// TIA Portal project "Urban Intersection Control System" (V17)

(* hardware
DEVICE "S7-1500/ET200MP station_1"  S7-1500 station
   slot 0: "Rail_0"  Rack  6ES7 590-1***0-0AA0
   slot 1: "PLC_UICS_01"  CPU 1512C-1 PN  6ES7 512-1CK00-0AB0  V2.9
      slot 3: "CPU display_1"  6ES7591-1AA00-0AA0
      slot 32768: "PROFINET interface_1"  X1
         slot 32769: "Port_1"  X1 P1
         slot 32770: "Port_2"  X1 P2
      slot 34817: "Virtual CP interface port_1"  Virtual CP interface port  Virtual CP interface port
DEVICE "HMI_1"  KTP1200 Basic PN
   slot 0: "HMI_1"  KTP1200 Basic PN  6AV2 123-2MB03-0AX0  17.0.0.0
   slot 1: "HMI_RT_1"  KTP1200 Basic PN  6AV2 123-2MB03-0AX0  17.0.0.0
   slot 5: "HMI_1.IE_CP_1"  PROFINET Interface  17.0.0.0
      slot 1: "PROFINET Interface_1"  PROFINET Interface
         slot 1: "Port_1"  Port
*)

// ===== PLC "PLC_UICS_01"  CPU 1512C-1 PN =====

VAR_GLOBAL   // PLC tag table "UICS_Table"
   "PB_Ped_Main_East" AT %I10.2 : Bool;   // Push button for pedestrian crossing on eastern Main Street
   "PB_Ped_Main_West" AT %I10.3 : Bool;   // Push button for pedestrian crossing on western Main Street
   "EM_Main_Override" AT %I10.6 : Bool;   // Emergency override signal (e.g. ambulances) on Main Street
   "EM_Cross_Override" AT %I10.7 : Bool;   // Emergency override signal on Cross Street
   "SENSOR_Main_Vehicle" AT %I11.0 : Bool;   // Vehicle detection sensor on Main Street
   "SENSOR_Cross_Vehicle" AT %I11.1 : Bool;   // Vehicle detection sensor on Cross Street
   "TL_Main_Red_West" AT %Q4.0 : Bool;   // Red traffic light signal for western Main Street
   "TL_Main_Yellow_West" AT %Q4.2 : Bool;   // Yellow traffic light signal for western Main Street
   "TL_Main_Green_West" AT %Q4.4 : Bool;   // Green traffic light signal for western Main Street
   "TL_Cross_Red_North" AT %Q4.6 : Bool;   // Red traffic light signal for northern Cross Street
   "TL_Cross_Yellow_North" AT %Q5.0 : Bool;   // Yellow traffic light signal for northern Cross Street
   "TL_Cross_Green_North" AT %Q5.2 : Bool;   // Green traffic light signal for northern Cross Street
   "PED_Main_Walk_West" AT %Q5.4 : Bool;   // Pedestrian walk signal for western Main Street
   "PED_Main_DontWalk_West" AT %Q5.6 : Bool;   // Pedestrian don’t-walk signal for western Main Street
   "PED_Cross_Walk_North" AT %Q6.0 : Bool;   // Pedestrian walk signal for northern Cross Street
   "PED_Cross_DontWalk_North" AT %Q6.2 : Bool;   // Pedestrian don’t-walk signal for northern Cross Street
   "PED_Warning_Buzzer" AT %Q6.4 : Bool;   // Audible alert for pedestrian crossing
   "SYS_Stop" AT %I10.1 : Bool;   // Emergency stop function
   "SYS_Start" AT %I10.0 : Bool;   // Begins the system
   "TL_Main_Red_East" AT %Q4.1 : Bool;   // Red traffic light signal for eastern Main Street
   "TL_Main_Yellow_East" AT %Q4.3 : Bool;   // Yellow traffic light signal for eastern Main Street
   "TL_Main_Green_East" AT %Q4.5 : Bool;   // Green traffic light signal for eastern Main Street
   "TL_Cross_Red_South" AT %Q4.7 : Bool;   // Red traffic light signal for southern Cross Street
   "TL_Cross_Yellow_South" AT %Q5.1 : Bool;   // Yellow traffic light signal for southern Cross Street
   "TL_Cross_Green_South" AT %Q5.3 : Bool;   // Green traffic light signal for southern Cross Street
   "PED_Main_Walk_East" AT %Q5.5 : Bool;   // Pedestrian walk signal for eastern Main Street
   "PED_Main_DontWalk_East" AT %Q5.7 : Bool;   // Pedestrian don’t-walk signal for eastern Main Street
   "PED_Cross_Walk_South" AT %Q6.1 : Bool;   // Pedestrian walk signal for southern Cross Street
   "PED_Cross_DontWalk_South" AT %Q6.3 : Bool;   // Pedestrian don’t-walk signal for southern Cross Street
   "PB_Ped_Cross_South" AT %I10.4 : Bool;   // Push button for pedestrian crossing on southern Cross Street
   "PB_Ped_Cross_North" AT %I10.5 : Bool;   // Push button for pedestrian crossing on northern Cross Street
   "PED_Main_Queue_East" AT %Q6.5 : Bool;   // Pedestrian queue signal for eastern Main Street
   "PED_Main_Queue_West" AT %Q6.6 : Bool;   // Pedestrian queue signal for western Main Street
   "PED_Cross_Queue_North" AT %Q6.7 : Bool;   // Pedestrian queue signal for southern Cross Street
   "PED_Cross_Queue_South" AT %Q7.0 : Bool;   // Pedestrian queue signal for northern Cross Street
END_VAR

DATA_BLOCK "Main_Control_System_DB"   // DB1
{ S7_Optimized_Access := 'TRUE' }
VERSION : 0.1
// stored: InstanceOfName Main_Control_System
"Main_Control_System"
BEGIN
END_DATA_BLOCK

DATA_BLOCK "Traffic_Light_Operations_DB"   // DB3
{ S7_Optimized_Access := 'TRUE' }
VERSION : 0.1
// stored: InstanceOfName Traffic_Light_Operations
"Traffic_Light_Operations"
BEGIN
END_DATA_BLOCK

DATA_BLOCK "Status_Reset_DB"   // DB7
{ S7_Optimized_Access := 'TRUE' }
VERSION : 0.1
// stored: InstanceOfName Status_Reset
"Status_Reset"
BEGIN
END_DATA_BLOCK

DATA_BLOCK "Pedestrian_Operations_DB"   // DB8
{ S7_Optimized_Access := 'TRUE' }
VERSION : 0.1
// stored: InstanceOfName Pedestrian_Operations
"Pedestrian_Operations"
BEGIN
END_DATA_BLOCK

DATA_BLOCK "Pedestrian_Crossing_DB"   // DB13
{ S7_Optimized_Access := 'TRUE' }
VERSION : 0.1
// stored: InstanceOfName Pedestrian_Crossing
"Pedestrian_Crossing"
BEGIN
END_DATA_BLOCK

// folder: System blocks/Program resources

DATA_BLOCK "MainStEast_Timer_DB"   // DB2
{ S7_Optimized_Access := 'TRUE' }
AUTHOR : Simatic
FAMILY : IEC
NAME : IEC_TMR
VERSION : 1.0
// stored: InstanceOfName IEC_TIMER
"IEC_TIMER"
BEGIN
END_DATA_BLOCK

DATA_BLOCK "CrossStNorth_Timer_DB"   // DB4
{ S7_Optimized_Access := 'TRUE' }
AUTHOR : Simatic
FAMILY : IEC
NAME : IEC_TMR
VERSION : 1.0
// stored: InstanceOfName IEC_TIMER
"IEC_TIMER"
BEGIN
END_DATA_BLOCK

DATA_BLOCK "CrossStSouth_Timer_DB"   // DB5
{ S7_Optimized_Access := 'TRUE' }
AUTHOR : Simatic
FAMILY : IEC
NAME : IEC_TMR
VERSION : 1.0
// stored: InstanceOfName IEC_TIMER
"IEC_TIMER"
BEGIN
END_DATA_BLOCK

DATA_BLOCK "MainStWest_Timer_DB"   // DB6
{ S7_Optimized_Access := 'TRUE' }
AUTHOR : Simatic
FAMILY : IEC
NAME : IEC_TMR
VERSION : 1.0
// stored: InstanceOfName IEC_TIMER
"IEC_TIMER"
BEGIN
END_DATA_BLOCK

DATA_BLOCK "Ped_MainStEast_Timer_DB"   // DB9
{ S7_Optimized_Access := 'TRUE' }
AUTHOR : Simatic
FAMILY : IEC
NAME : IEC_TMR
VERSION : 1.0
// stored: InstanceOfName IEC_TIMER
"IEC_TIMER"
BEGIN
END_DATA_BLOCK

DATA_BLOCK "Ped_MainStWest_Timer_DB"   // DB10
{ S7_Optimized_Access := 'TRUE' }
AUTHOR : Simatic
FAMILY : IEC
NAME : IEC_TMR
VERSION : 1.0
// stored: InstanceOfName IEC_TIMER
"IEC_TIMER"
BEGIN
END_DATA_BLOCK

DATA_BLOCK "Ped_CrossStSouth_Timer_DB"   // DB11
{ S7_Optimized_Access := 'TRUE' }
AUTHOR : Simatic
FAMILY : IEC
NAME : IEC_TMR
VERSION : 1.0
// stored: InstanceOfName IEC_TIMER
"IEC_TIMER"
BEGIN
END_DATA_BLOCK

DATA_BLOCK "Ped_CrossStNorth_Timer_DB"   // DB12
{ S7_Optimized_Access := 'TRUE' }
AUTHOR : Simatic
FAMILY : IEC
NAME : IEC_TMR
VERSION : 1.0
// stored: InstanceOfName IEC_TIMER
"IEC_TIMER"
BEGIN
END_DATA_BLOCK

// folder: (top level)

FUNCTION_BLOCK "Main_Control_System"   // FB1, LAD
{ S7_Optimized_Access := 'TRUE' }
VERSION : 0.1
   VAR_INPUT
      System_Start : Bool;   // Activates the system
      System_Stop : Bool;   // Emergency stop function
   END_VAR
   VAR
      System_Latch : Bool;   // Allows the system to remain active after initially starting up
      System_Running : Bool;   // System is actively running
      Emergency_Stop : Bool;   // Emergency stop activated flag
      HMI_Start_Command : Bool;   // Allows HMI to start the system
      HMI_Stop_Command : Bool;   // Allows HMI to stop the system
      HMI_Latch_Command : Bool;   // Allows HMI visualization to remain active after initially starting up
      HMI_Run_Command : Bool;   // Allows HMI to run the system
   END_VAR
BEGIN

REGION Network 1: System Start
   // Starts the system if all conditions are met
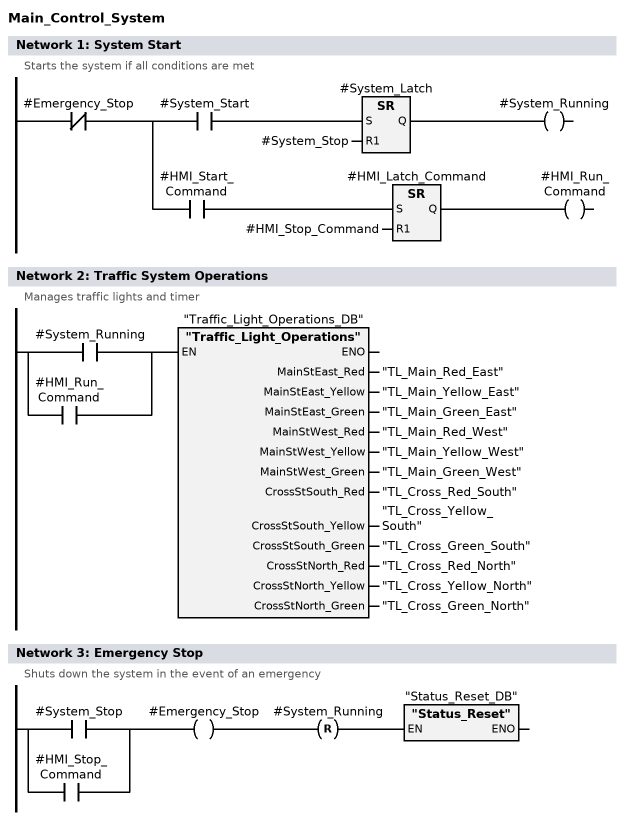
   RUNG wire#powerrail
      I_Contact( #Emergency_Stop )
      wire#w1
      Contact( #System_Start )
      S_SR(operand := #System_Latch, r1 := #System_Stop)
      Coil( #System_Running )
   END_RUNG
   RUNG wire#w1
      Contact( #HMI_Start_Command )
      S_SR(operand := #HMI_Latch_Command, r1 := #HMI_Stop_Command)
      Coil( #HMI_Run_Command )
   END_RUNG
   // the same network as SCL:
   IF NOT #Emergency_Stop AND #System_Start THEN
       #System_Latch := TRUE;   // SR flip-flop
   END_IF;
   IF #System_Stop THEN #System_Latch := FALSE; END_IF;
   #System_Running := #System_Latch;
   IF NOT #Emergency_Stop AND #HMI_Start_Command THEN
       #HMI_Latch_Command := TRUE;   // SR flip-flop
   END_IF;
   IF #HMI_Stop_Command THEN #HMI_Latch_Command := FALSE; END_IF;
   #HMI_Run_Command := #HMI_Latch_Command;
END_REGION

REGION Network 2: Traffic System Operations
   // Manages traffic lights and timer
   RUNG wire#powerrail
      Contact( #System_Running )
      wire#w1
      "Traffic_Light_Operations_DB"(MainStEast_Red => "TL_Main_Red_East", MainStEast_Yellow => "TL_Main_Yellow_East", MainStEast_Green => "TL_Main_Green_East", MainStWest_Red => "TL_Main_Red_West", MainStWest_Yellow => "TL_Main_Yellow_West", MainStWest_Green => "TL_Main_Green_West", CrossStSouth_Red => "TL_Cross_Red_South", CrossStSouth_Yellow => "TL_Cross_Yellow_South", CrossStSouth_Green => "TL_Cross_Green_South", CrossStNorth_Red => "TL_Cross_Red_North", CrossStNorth_Yellow => "TL_Cross_Yellow_North", CrossStNorth_Green => "TL_Cross_Green_North")
   END_RUNG
   RUNG wire#powerrail
      Contact( #HMI_Run_Command )
   END_RUNG wire#w1
   // the same network as SCL:
   IF #System_Running OR #HMI_Run_Command THEN
       "Traffic_Light_Operations_DB"(MainStEast_Red => "TL_Main_Red_East",   // "Traffic_Light_Operations"
                               MainStEast_Yellow => "TL_Main_Yellow_East",
                               MainStEast_Green => "TL_Main_Green_East",
                               MainStWest_Red => "TL_Main_Red_West",
                               MainStWest_Yellow => "TL_Main_Yellow_West",
                               MainStWest_Green => "TL_Main_Green_West",
                               CrossStSouth_Red => "TL_Cross_Red_South",
                               CrossStSouth_Yellow => "TL_Cross_Yellow_South",
                               CrossStSouth_Green => "TL_Cross_Green_South",
                               CrossStNorth_Red => "TL_Cross_Red_North",
                               CrossStNorth_Yellow => "TL_Cross_Yellow_North",
                               CrossStNorth_Green => "TL_Cross_Green_North");
   END_IF;
END_REGION

REGION Network 3: Emergency Stop
   // Shuts down the system in the event of an emergency
   RUNG wire#powerrail
      Contact( #System_Stop )
      wire#w1
      Coil( #Emergency_Stop )
      R_Coil( #System_Running )
      "Status_Reset_DB"()
   END_RUNG
   RUNG wire#powerrail
      Contact( #HMI_Stop_Command )
   END_RUNG wire#w1
   // the same network as SCL:
   #Emergency_Stop := #System_Stop OR #HMI_Stop_Command;
   IF #Emergency_Stop THEN
       #System_Running := FALSE;
       "Status_Reset_DB"();   // "Status_Reset"
   END_IF;
END_REGION
END_FUNCTION_BLOCK

FUNCTION_BLOCK "Traffic_Light_Operations"   // FB2, LAD
{ S7_Optimized_Access := 'TRUE' }
VERSION : 0.1
   VAR_OUTPUT
      MainStEast_Red : Bool;   // Red traffic light signal for eastern Main Street
      MainStEast_Yellow : Bool;   // Yellow traffic light signal for eastern Main Street
      MainStEast_Green : Bool;   // Green traffic light signal for eastern Main Street
      MainStWest_Red : Bool;   // Red traffic light signal for western Main Street
      MainStWest_Yellow : Bool;   // Yellow traffic light signal for western Main Street
      MainStWest_Green : Bool;   // Green traffic light signal for western Main Street
      CrossStSouth_Red : Bool;   // Red traffic light signal for southern Cross Street
      CrossStSouth_Yellow : Bool;   // Yellow traffic light signal for southern Cross Street
      CrossStSouth_Green : Bool;   // Green traffic light signal for southern Cross Street
      CrossStNorth_Red : Bool;   // Red traffic light signal for northern Cross Street
      CrossStNorth_Yellow : Bool;   // Yellow traffic light signal for northern Cross Street
      CrossStNorth_Green : Bool;   // Green traffic light signal for northern Cross Street
   END_VAR
   VAR
      Traffic_Operations_Step : Int;   // Controls the state of traffic operations
      MainStEast_Seconds : Int;   // Allows HMI to read eastern Main Street traffic time
      MainStWest_Seconds : Int;   // Allows HMI to read western Main Street traffic time
      CrossStNorth_Seconds : Int;   // Allows HMI to read northern Cross Street traffic time
      CrossStSouth_Seconds : Int;   // Allows HMI to read southern Cross Street traffic time
      Initialize_Operation : Bool;   // Initiates traffic operations
   END_VAR
   VAR_TEMP
      MainStEast_ET_DInt : DInt;
      MainStEast_ET_Div : DInt;
      CrossStSouth_ET_DInt : DInt;
      CrossStSouth_ET_Div : DInt;
      MainStWest_ET_DInt : DInt;
      MainStWest_ET_Div : DInt;
      CrossStNorth_ET_DInt : DInt;
      CrossStNorth_ET_Div : DInt;
   END_VAR
   VAR_TEMP   // added for the SCL form of the ladder/FBD networks
      _w1 : Bool;
   END_VAR
BEGIN

REGION Network 1: Red Light Control
   // Organization of red traffic lights for Main Street and Cross Street
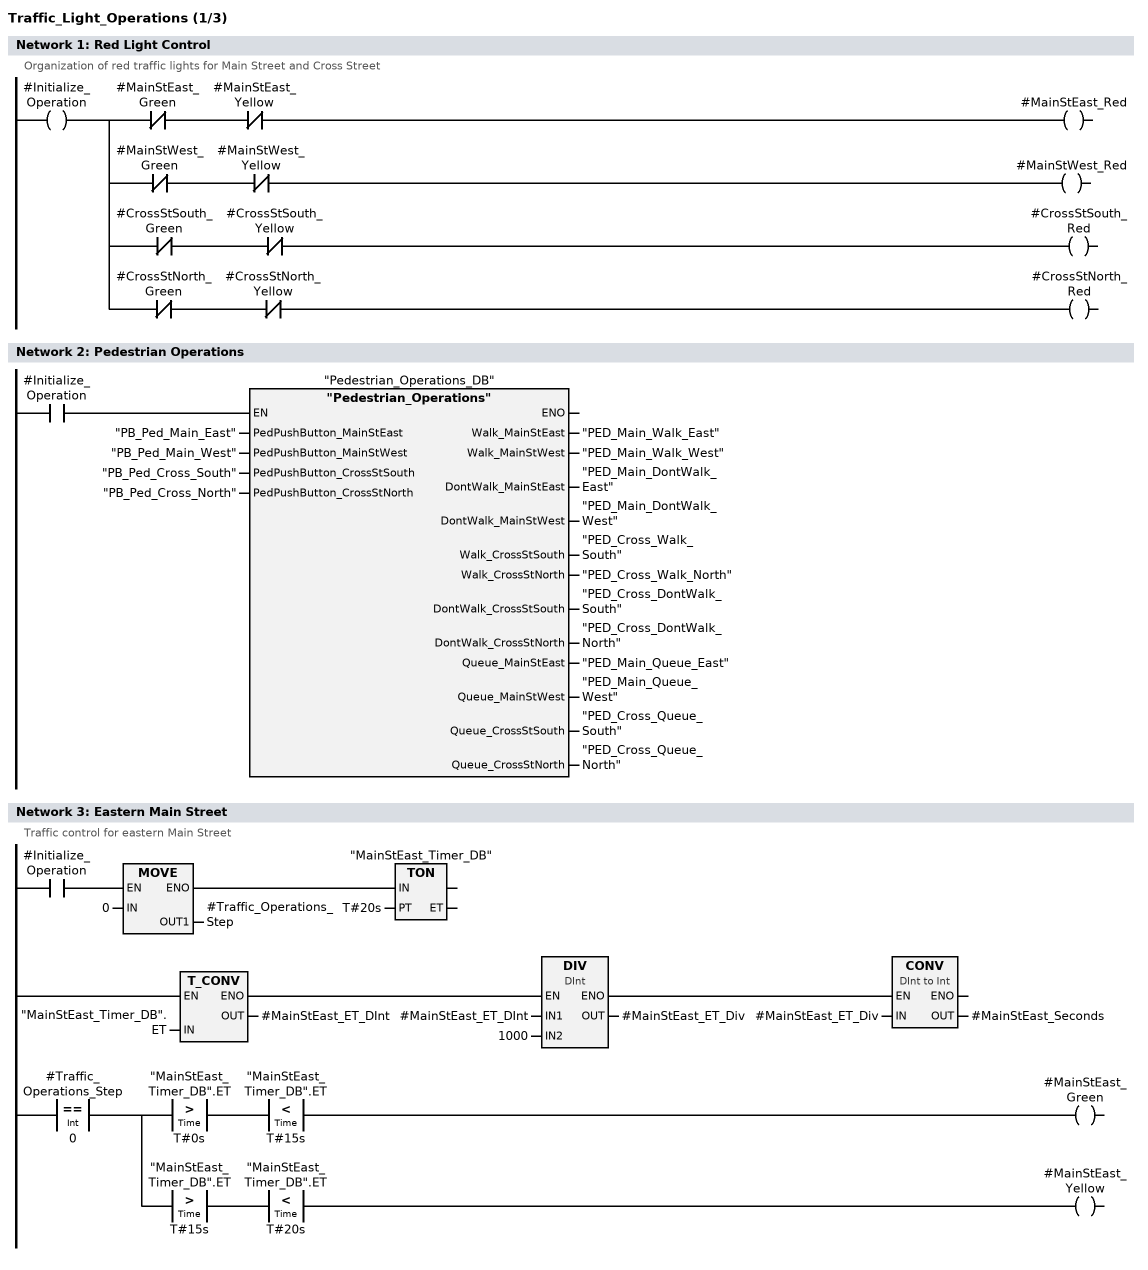
   RUNG wire#powerrail
      Coil( #Initialize_Operation )
      wire#w1
      I_Contact( #MainStEast_Green )
      I_Contact( #MainStEast_Yellow )
      Coil( #MainStEast_Red )
   END_RUNG
   RUNG wire#w1
      I_Contact( #MainStWest_Green )
      I_Contact( #MainStWest_Yellow )
      Coil( #MainStWest_Red )
   END_RUNG
   RUNG wire#w1
      I_Contact( #CrossStSouth_Green )
      I_Contact( #CrossStSouth_Yellow )
      Coil( #CrossStSouth_Red )
   END_RUNG
   RUNG wire#w1
      I_Contact( #CrossStNorth_Green )
      I_Contact( #CrossStNorth_Yellow )
      Coil( #CrossStNorth_Red )
   END_RUNG
   // the same network as SCL:
   #Initialize_Operation := TRUE;
   #MainStEast_Red := NOT #MainStEast_Green AND NOT #MainStEast_Yellow;
   #MainStWest_Red := NOT #MainStWest_Green AND NOT #MainStWest_Yellow;
   #CrossStSouth_Red := NOT #CrossStSouth_Green AND NOT #CrossStSouth_Yellow;
   #CrossStNorth_Red := NOT #CrossStNorth_Green AND NOT #CrossStNorth_Yellow;
END_REGION

REGION Network 2: Pedestrian Operations
   RUNG wire#powerrail
      Contact( #Initialize_Operation )
      "Pedestrian_Operations_DB"(PedPushButton_MainStEast := "PB_Ped_Main_East", PedPushButton_MainStWest := "PB_Ped_Main_West", PedPushButton_CrossStSouth := "PB_Ped_Cross_South", PedPushButton_CrossStNorth := "PB_Ped_Cross_North", Walk_MainStEast => "PED_Main_Walk_East", Walk_MainStWest => "PED_Main_Walk_West", DontWalk_MainStEast => "PED_Main_DontWalk_East", DontWalk_MainStWest => "PED_Main_DontWalk_West", Walk_CrossStSouth => "PED_Cross_Walk_South", Walk_CrossStNorth => "PED_Cross_Walk_North", DontWalk_CrossStSouth => "PED_Cross_DontWalk_South", DontWalk_CrossStNorth => "PED_Cross_DontWalk_North", Queue_MainStEast => "PED_Main_Queue_East", Queue_MainStWest => "PED_Main_Queue_West", Queue_CrossStSouth => "PED_Cross_Queue_South", Queue_CrossStNorth => "PED_Cross_Queue_North")
   END_RUNG
   // the same network as SCL:
   IF #Initialize_Operation THEN
       "Pedestrian_Operations_DB"(PedPushButton_MainStEast := "PB_Ped_Main_East",   // "Pedestrian_Operations"
                               PedPushButton_MainStWest := "PB_Ped_Main_West",
                               PedPushButton_CrossStSouth := "PB_Ped_Cross_South",
                               PedPushButton_CrossStNorth := "PB_Ped_Cross_North",
                               Walk_MainStEast => "PED_Main_Walk_East",
                               Walk_MainStWest => "PED_Main_Walk_West",
                               DontWalk_MainStEast => "PED_Main_DontWalk_East",
                               DontWalk_MainStWest => "PED_Main_DontWalk_West",
                               Walk_CrossStSouth => "PED_Cross_Walk_South",
                               Walk_CrossStNorth => "PED_Cross_Walk_North",
                               DontWalk_CrossStSouth => "PED_Cross_DontWalk_South",
                               DontWalk_CrossStNorth => "PED_Cross_DontWalk_North",
                               Queue_MainStEast => "PED_Main_Queue_East",
                               Queue_MainStWest => "PED_Main_Queue_West",
                               Queue_CrossStSouth => "PED_Cross_Queue_South",
                               Queue_CrossStNorth => "PED_Cross_Queue_North");
   END_IF;
END_REGION

REGION Network 3: Eastern Main Street
   // Traffic control for eastern Main Street
   // ENO of a box is taken as its EN; it also drops when the box reports an error
   IF #Initialize_Operation THEN #Traffic_Operations_Step := 0; END_IF;
   "MainStEast_Timer_DB".TON(IN := #Initialize_Operation, PT := T#20s);
   #MainStEast_ET_DInt := T_CONV(IN := "MainStEast_Timer_DB".ET);
   #MainStEast_ET_Div := #MainStEast_ET_DInt / 1000;
   #MainStEast_Seconds := DINT_TO_INT(#MainStEast_ET_Div);
   #_w1 := #Traffic_Operations_Step = 0;
   #MainStEast_Green := #_w1 AND ("MainStEast_Timer_DB".ET > T#0s) AND ("MainStEast_Timer_DB".ET < T#15s);
   #MainStEast_Yellow := #_w1 AND ("MainStEast_Timer_DB".ET > T#15s) AND ("MainStEast_Timer_DB".ET < T#20s);
END_REGION

REGION Network 4: Western Main Street
   // Traffic control for western Main Street
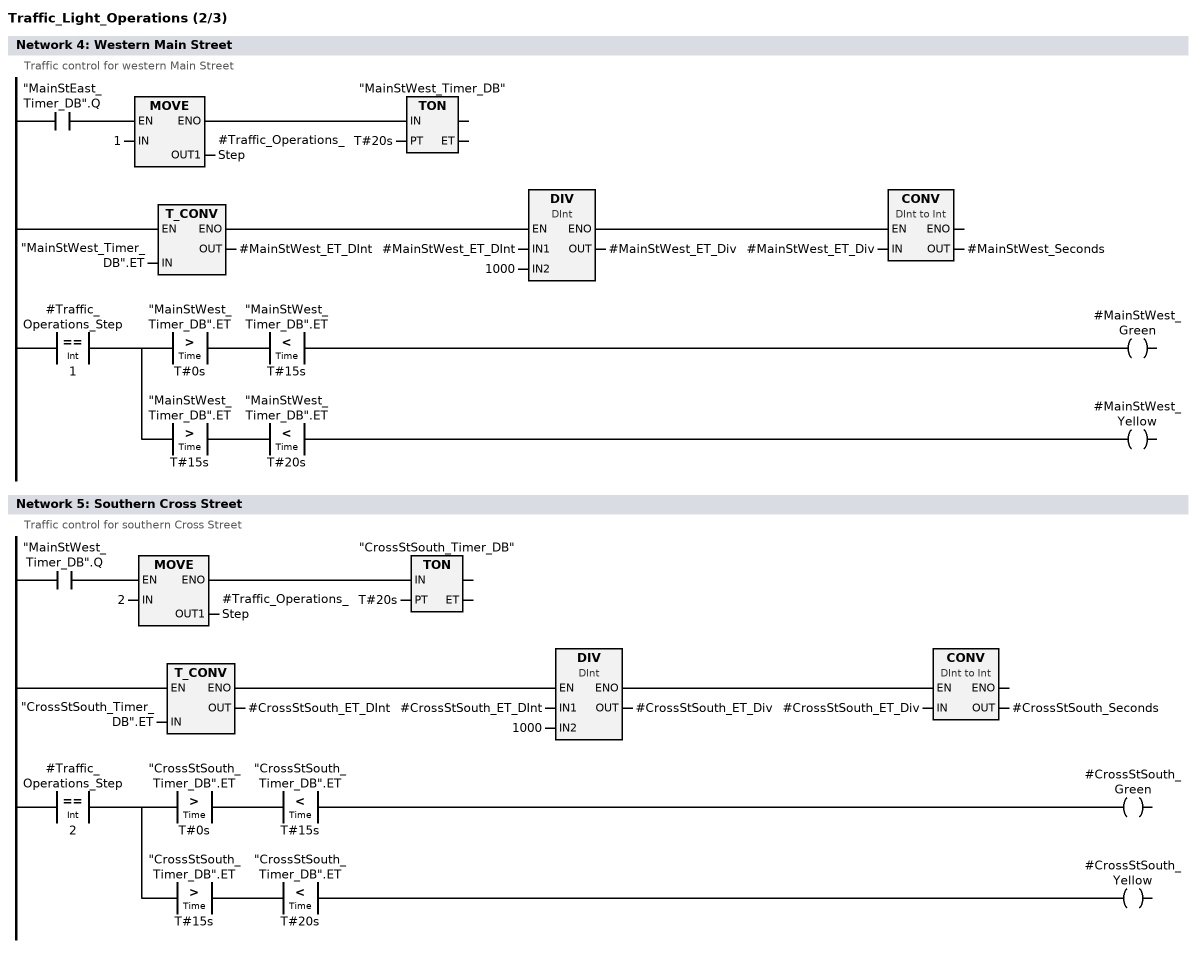
   // ENO of a box is taken as its EN; it also drops when the box reports an error
   IF "MainStEast_Timer_DB".Q THEN #Traffic_Operations_Step := 1; END_IF;
   "MainStWest_Timer_DB".TON(IN := "MainStEast_Timer_DB".Q, PT := T#20s);
   #MainStWest_ET_DInt := T_CONV(IN := "MainStWest_Timer_DB".ET);
   #MainStWest_ET_Div := #MainStWest_ET_DInt / 1000;
   #MainStWest_Seconds := DINT_TO_INT(#MainStWest_ET_Div);
   #_w1 := #Traffic_Operations_Step = 1;
   #MainStWest_Green := #_w1 AND ("MainStWest_Timer_DB".ET > T#0s) AND ("MainStWest_Timer_DB".ET < T#15s);
   #MainStWest_Yellow := #_w1 AND ("MainStWest_Timer_DB".ET > T#15s) AND ("MainStWest_Timer_DB".ET < T#20s);
END_REGION

REGION Network 5: Southern Cross Street
   // Traffic control for southern Cross Street
   // ENO of a box is taken as its EN; it also drops when the box reports an error
   IF "MainStWest_Timer_DB".Q THEN #Traffic_Operations_Step := 2; END_IF;
   "CrossStSouth_Timer_DB".TON(IN := "MainStWest_Timer_DB".Q, PT := T#20s);
   #CrossStSouth_ET_DInt := T_CONV(IN := "CrossStSouth_Timer_DB".ET);
   #CrossStSouth_ET_Div := #CrossStSouth_ET_DInt / 1000;
   #CrossStSouth_Seconds := DINT_TO_INT(#CrossStSouth_ET_Div);
   #_w1 := #Traffic_Operations_Step = 2;
   #CrossStSouth_Green := #_w1 AND ("CrossStSouth_Timer_DB".ET > T#0s) AND ("CrossStSouth_Timer_DB".ET < T#15s);
   #CrossStSouth_Yellow := #_w1 AND ("CrossStSouth_Timer_DB".ET > T#15s) AND ("CrossStSouth_Timer_DB".ET < T#20s);
END_REGION

REGION Network 6: Northern Cross Street
   // Traffic control for northern Cross Street
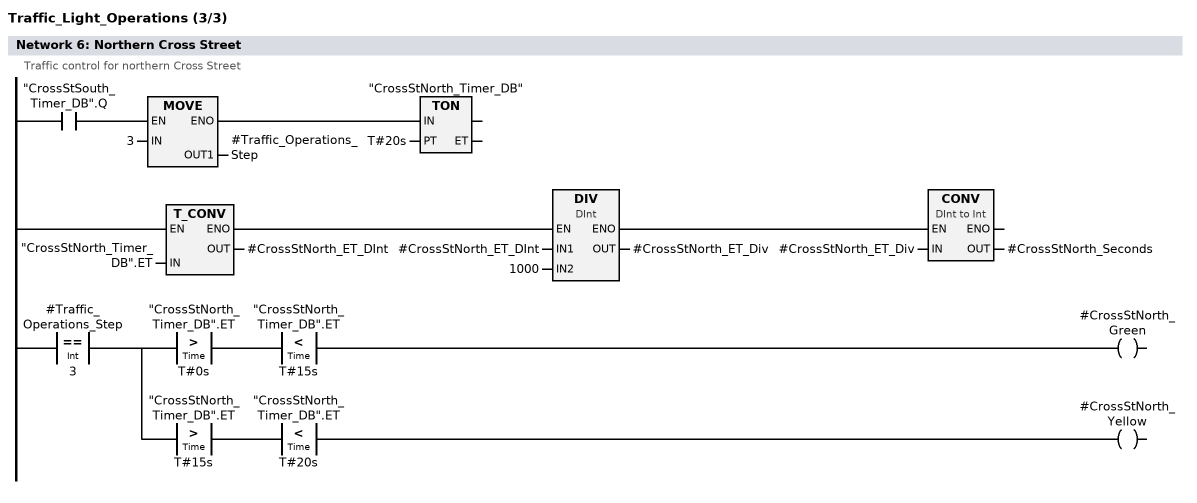
   // ENO of a box is taken as its EN; it also drops when the box reports an error
   IF "CrossStSouth_Timer_DB".Q THEN #Traffic_Operations_Step := 3; END_IF;
   "CrossStNorth_Timer_DB".TON(IN := "CrossStSouth_Timer_DB".Q, PT := T#20s);
   #CrossStNorth_ET_DInt := T_CONV(IN := "CrossStNorth_Timer_DB".ET);
   #CrossStNorth_ET_Div := #CrossStNorth_ET_DInt / 1000;
   #CrossStNorth_Seconds := DINT_TO_INT(#CrossStNorth_ET_Div);
   #_w1 := #Traffic_Operations_Step = 3;
   #CrossStNorth_Green := #_w1 AND ("CrossStNorth_Timer_DB".ET > T#0s) AND ("CrossStNorth_Timer_DB".ET < T#15s);
   #CrossStNorth_Yellow := #_w1 AND ("CrossStNorth_Timer_DB".ET > T#15s) AND ("CrossStNorth_Timer_DB".ET < T#20s);
END_REGION
END_FUNCTION_BLOCK

FUNCTION_BLOCK "Status_Reset"   // FB3, LAD
{ S7_Optimized_Access := 'TRUE' }
VERSION : 0.1
BEGIN

REGION Network 1: Traffic Status Reset
   // Resets the status of the traffic timers, traffic lights, and other variables
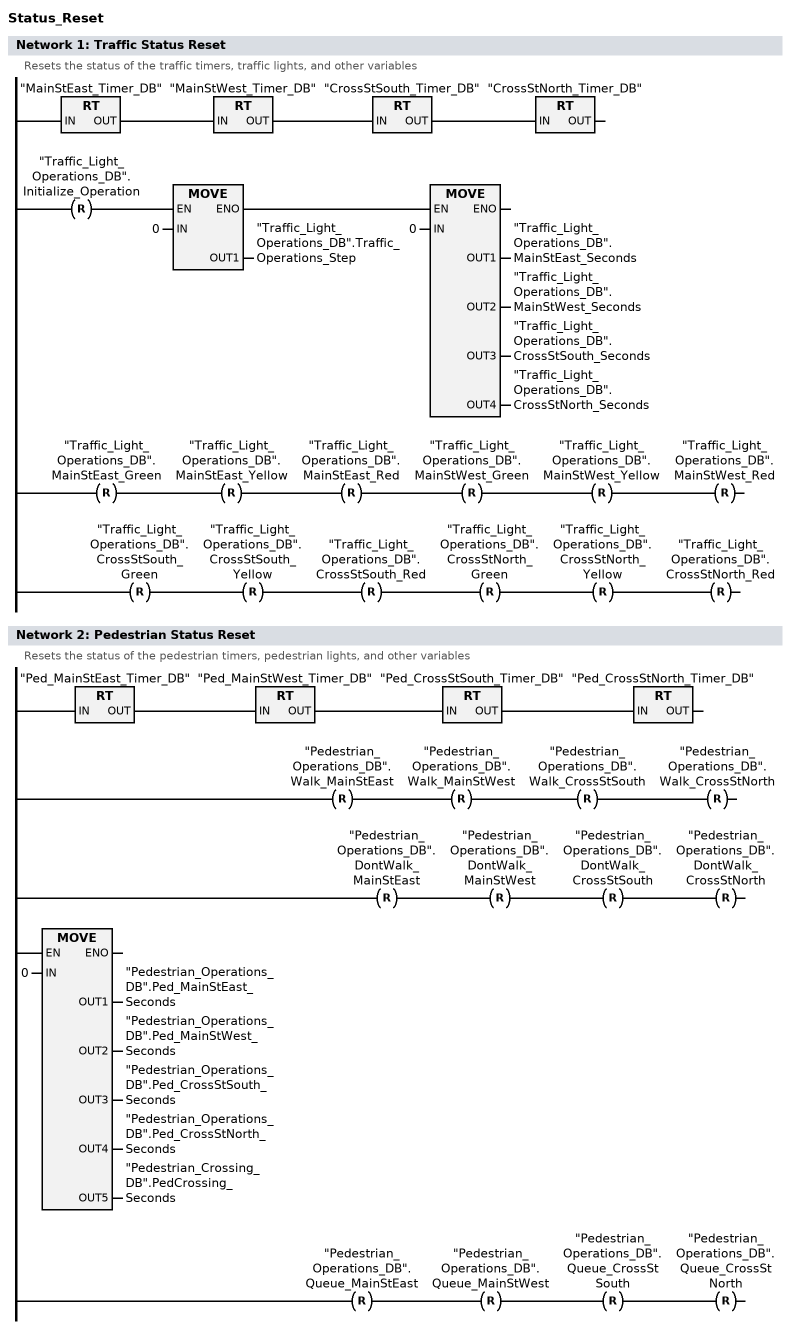
   RUNG wire#powerrail
      RT_Coil( "MainStEast_Timer_DB" )
      RT_Coil( "MainStWest_Timer_DB" )
      RT_Coil( "CrossStSouth_Timer_DB" )
      RT_Coil( "CrossStNorth_Timer_DB" )
   END_RUNG
   RUNG wire#powerrail
      R_Coil( "Traffic_Light_Operations_DB".Initialize_Operation )
      Move(in := 0, out1 => "Traffic_Light_Operations_DB".Traffic_Operations_Step)
      Move(in := 0, out1 => "Traffic_Light_Operations_DB".MainStEast_Seconds, out2 => "Traffic_Light_Operations_DB".MainStWest_Seconds, out3 => "Traffic_Light_Operations_DB".CrossStSouth_Seconds, out4 => "Traffic_Light_Operations_DB".CrossStNorth_Seconds)
   END_RUNG
   RUNG wire#powerrail
      R_Coil( "Traffic_Light_Operations_DB".MainStEast_Green )
      R_Coil( "Traffic_Light_Operations_DB".MainStEast_Yellow )
      R_Coil( "Traffic_Light_Operations_DB".MainStEast_Red )